        [28]   // FV26 Chill Down Pressure
        [29]   // FV26 Chill Down Current Time
        [2]   // FV26 Level Probes
        [30]   // FV26 Time since Clean
        [32]   // FV26 CIP Selected
        [32].0   // FV26 Request Channel 1 CIP
        [32].1   // FV26 Request Channel 2 CIP
        [33]   // FV26 Rotocheck
        [33].0   // FV26 Enable Rotocheck
        [33].1   // FV26 Rotocheck Fault
        [38]   // FV26 Pressure Difference Bottom-Top (psi)
        [39]   // FV26 Pressure Difference Calibration Offset
        [3]   // FV26 Top Pressure Status
        [40]   // FV26 Cropping Status 0=Not Done 1=Running 2=Done 3=Done+48hrs
        [43]   // FV26 Hours since Yeast Cropping
        [4]   // FV26 Yeast Status
        [50]   // FV26 FiltrateReturnStatus 0=Not Done 1=Running 2=Done
        [5]   // FV26 Aging Status
        [60].3   // FV26 Top Pressure Chill Down
        [6]   // FV26 Valve Routes
        [6].0   // FV26 Inlet Main to Drain Open
        [6].1   // FV26 Filling Valve Not Closed
        [6].2   // FV26 Filling Inlet Open
        [6].3   // FV26 Bypass Route Open Open
        [6].4   // FV26 Green Beer Open
        [6].5   // FV26 Yeast Removal Open
        [6].6   // FV26 Filtrate Open
        [6].7   // FV26 CIP Open
        [7]   // FV26 Top Pressure Control Actual Pressure
        [7].0   // FV26 Yeast Status Filtrate Return
        [8]   // FV26 Log Message
        [9]   // FV26 Item Fault
   FR_N27 : INT[265] := ([0] := 227, [1] := 3, [3] := 2, [5] := 4, [6] := 8, [7] := 1030, [8] := 12227, [9] := -1, [10] := 2387, [11] := 9672, [12] := 1575, [13] := 2902, [14] := 603, [15] := 1292, [16] := 891, [17] := 9083, [18] := 12, [19] := 8975, [20] := 1, [21] := 4, [22] := 1000, [23] := 50, [24] := 1050, [25] := 950, [26] := 1000, [27] := 8, [30] := 2, [33] := 1, [37] := 702, [38] := 1357, [39] := 65, [52] := 1, [60] := 4, [68] := 5311, [69] := 172, [90] := 1, [91] := 251, [92] := 841, [100] := 43, [101] := 49, [102] := 55, [103] := 13, [104] := 14, [105] := 15, [106] := 16, [107] := 17, [108] := 97, [109] := -1, [110] := -1, [111] := -1, [112] := -1, [113] := -1, [114] := -1, [115] := -1, [116] := -1, [117] := -1, [118] := -1, [119] := -1, [120] := -1, [121] := -1,
        [122] := -1, [123] := -1, [124] := -1, [125] := -1, [126] := -1, [127] := -1, [128] := -1, [129] := -1, [130] := -1, [131] := -1, [132] := -1, [133] := -1, [134] := -1, [135] := -1, [136] := -1, [137] := -1, [138] := -1, [139] := -1, [140] := -1, [141] := -1, [142] := -1, [143] := -1, [144] := -1, [145] := -1, [146] := -1, [147] := -1, [148] := -1, [149] := -1);   // FV27
        [0]   // FV27
        [100]   // FV27 Checklist Data
        [10]   // FV27 Bottom Pressure
        [11]   // FV27 Damped Level
        [12]   // FV27 Cone Radius
        [13]   // FV27 Cone Height
        [14]   // FV27 Volume (HL)
        [19]   // FV27 Height above LTX
        [1]   // FV27 Status 0=Clean,1=Fill,2=Par t,3=Ferment,4=?,5=?, 6=?,7=?,8=Emptying,9 =Dirty,10-13=CIP
        [20]   // FV27 Top Pressure Bits
        [20].2   // FV27 Top Pressure Chill Down
        [20].5   // FV27 Top Pressure Step Channel 1 CIP
        [20].6   // FV27 Top Pressure Bits Ch1 CIP Complete
        [20].7   // FV27 Top Pressure Step Channel 2 CIP
        [20].8   // FV27 Top Pressure Bits Ch2 CIP Complete
        [21]   // FV27 Top Pressure Step Flags
        [21].0   // FV27 Top Pressure Control Over Pressure
        [21].4   // FV27 Top Pressure Open Vent
        [21].5   // FV27 Top Pressure Control Open Vent Actuator
        [21].6   // FV27 Over Top Pressure Limit
        [21].8   // FV27 Top Pressure Control Over Pressure Alarm
        [22]   // FV27 Top Pressure Setpoint
        [23]   // FV27 Top Pressure Deadband
        [24]   // FV27 Top Pressure Upper Limit
        [25]   // FV27 Top Pressure Lower Limit
        [26]   // FV27 Fermenting Pressure
        [27]   // FV27 Chill Down Time
        [28]   // FV27 Chill Down Pressure
        [29]   // FV27 Chill Down Current Time
        [2]   // FV27 Level Probes
        [30]   // FV27 Time since Clean
        [32]   // FV27 CIP Selected
        [32].0   // FV27 Request Channel 1 CIP
        [32].1   // FV27 Request Channel 2 CIP
        [33]   // FV27 Rotocheck
        [33].0   // FV27 Enable Rotocheck
        [33].1   // FV27 Rotocheck Fault
        [38]   // FV27 Pressure Difference Bottom-Top (psi)
        [39]   // FV27 Pressure Difference Calibration Offset
        [3]   // FV27 Top Pressure Status
        [40]   // FV27 Cropping Status 0=Not Done 1=Running 2=Done 3=Done+48hrs
        [43]   // FV27 Hours since Yeast Cropping
        [4]   // FV27 Yeast Status
        [50]   // FV27 FiltrateReturnStatus 0=Not Done 1=Running 2=Done
        [5]   // FV27 Aging Status
        [60].3   // FV27 Top Pressure Chill Down
        [6]   // FV27 Valve Routes
        [6].0   // FV27 Inlet Main to Drain Open
        [6].1   // FV27 Filling Valve Not Closed
        [6].2   // FV27 Filling Inlet Open
        [6].3   // FV27 Bypass Route Open Open
        [6].4   // FV27 Green Beer Open
        [6].5   // FV27 Yeast Removal Open
        [6].6   // FV27 Filtrate Open
        [6].7   // FV27 CIP Open
        [7]   // FV27 Top Pressure Control Actual Pressure
        [7].0   // FV27 Yeast Status Filtrate Return
        [8]   // FV27 Log Message
        [90]   // Vent Actuations Counter
        [91]   // FV27/PTX01 FV27 top pressure minimum
        [92]   // FV27/PTX01 FV27 top pressure maximum
        [9]   // FV27 Item Fault
   FR_N28 : INT[265] := ([0] := 228, [1] := 3, [2] := 1, [3] := 4, [4] := 30, [5] := 6, [6] := 8, [7] := 1, [8] := 12228, [9] := -1, [10] := 1150, [11] := 8680, [12] := 1575, [13] := 2902, [14] := 526, [15] := 1149, [16] := 792, [17] := 8073, [18] := 12, [19] := 7977, [20] := 1, [21] := 18, [22] := 167, [24] := 167, [25] := 167, [26] := 1000, [27] := 12, [29] := 10, [30] := 23, [33] := 1, [37] := 702, [38] := 1149, [52] := 1, [60] := 16, [68] := 5228, [69] := 5228, [100] := 47, [101] := 53, [102] := 59, [103] := 27, [104] := 28, [105] := 29, [106] := 30, [107] := 31, [108] := 98, [109] := -1, [110] := -1, [111] := -1, [112] := -1, [113] := -1, [114] := -1, [115] := -1, [116] := -1, [117] := -1, [118] := -1, [119] := -1, [120] := -1, [121] := -1, [122] := -1, [123] := -1,
        [124] := -1, [125] := -1, [126] := -1, [127] := -1, [128] := -1, [129] := -1, [130] := -1, [131] := -1, [132] := -1, [133] := -1, [134] := -1, [135] := -1, [136] := -1, [137] := -1, [138] := -1, [139] := -1, [140] := -1, [141] := -1, [142] := -1, [143] := -1, [144] := -1, [145] := -1, [146] := -1, [147] := -1, [148] := -1, [149] := -1);   // FV28
        [0]   // FV28
        [100]   // FV28 Checklist Data
        [10]   // FV28 Bottom Pressure
        [11]   // FV28 Damped Level
        [12]   // FV28 Cone Radius
        [13]   // FV28 Cone Height
        [14]   // FV28 Volume (HL)
        [19]   // FV28 Height above LTX
        [1]   // FV28 Status 0=Clean,1=Fill,2=Par t,3=Ferment,4=?,5=?, 6=?,7=?,8=Emptying,9 =Dirty,10-13=CIP
        [20]   // FV28 Top Pressure Bits
        [20].2   // FV28 Top Pressure Chill Down
        [20].5   // FV28 Top Pressure Step Channel 1 CIP
        [20].6   // FV28 Top Pressure Bits Ch1 CIP Complete
        [20].7   // FV28 Top Pressure Step Channel 2 CIP
        [20].8   // FV28 Top Pressure Bits Ch2 CIP Complete
        [21]   // FV28 Top Pressure Step Flags
        [21].0   // FV28 Top Pressure Control Over Pressure
        [21].4   // FV28 Top Pressure Open Vent
        [21].5   // FV28 Top Pressure Control Open Vent Actuator
        [21].6   // FV28 Over Top Pressure Limit
        [21].8   // FV28 Top Pressure Control Over Pressure Alarm
        [22]   // FV28 Top Pressure Setpoint
        [23]   // FV28 Top Pressure Deadband
        [24]   // FV28 Top Pressure Upper Limit
        [25]   // FV28 Top Pressure Lower Limit
        [26]   // FV28 Fermenting Pressure
        [27]   // FV28 Chill Down Time
        [28]   // FV28 Chill Down Pressure
        [29]   // FV28 Chill Down Current Time
        [2]   // FV28 Level Probes
        [30]   // FV28 Time since Clean
        [32]   // FV28 CIP Selected
        [32].0   // FV28 Request Channel 1 CIP
        [32].1   // FV28 Request Channel 2 CIP
        [33]   // FV28 Rotocheck
        [33].0   // FV28 Enable Rotocheck
        [33].1   // FV28 Rotocheck Fault
        [38]   // FV28 Pressure Difference Bottom-Top (psi)
        [39]   // FV28 Pressure Difference Calibration Offset
        [3]   // FV28 Top Pressure Status
        [40]   // FV28 Cropping Status 0=Not Done 1=Running 2=Done 3=Done+48hrs
        [43]   // FV28 Hours since Yeast Cropping
        [4]   // FV28 Yeast Status
        [50]   // FV28 FiltrateReturnStatus 0=Not Done 1=Running 2=Done
        [5]   // FV28 Aging Status
        [60].3   // FV28 Top Pressure Chill Down
        [6]   // FV28 Valve Routes
        [6].0   // FV28 Inlet Main to Drain Open
        [6].1   // FV28 Filling Valve Not Closed
        [6].2   // FV28 Filling Inlet Open
        [6].3   // FV28 Bypass Route Open Open
        [6].4   // FV28 Green Beer Open
        [6].5   // FV28 Yeast Removal Open
        [6].6   // FV28 Filtrate Open
        [6].7   // FV28 CIP Open
        [7]   // FV28 Top Pressure Control Actual Pressure
        [7].0   // FV28 Yeast Status Filtrate Return
        [8]   // FV28 Log Message
        [9]   // FV28 Item Fault
   FR_N29 : INT[265] := ([0] := 229, [1] := 9, [2] := 2, [3] := 6, [4] := 2, [6] := 8, [7] := 6, [8] := 12229, [9] := -1, [10] := -1, [11] := -50, [12] := 1575, [13] := 2902, [15] := -7, [16] := -5, [17] := -51, [18] := 12, [19] := -50, [20] := 1, [21] := 33, [22] := -125, [23] := 50, [24] := -75, [25] := -175, [26] := 1000, [27] := 8, [30] := 39, [33] := 1, [37] := 702, [38] := -7, [52] := 1, [60] := 64, [69] := 5213, [100] := 46, [101] := 52, [102] := 58, [103] := 32, [104] := 33, [105] := 34, [106] := 35, [107] := 36, [108] := 99, [109] := -1, [110] := -1, [111] := -1, [112] := -1, [113] := -1, [114] := -1, [115] := -1, [116] := -1, [117] := -1, [118] := -1, [119] := -1, [120] := -1, [121] := -1, [122] := -1, [123] := -1, [124] := -1, [125] := -1, [126] := -1,
        [127] := -1, [128] := -1, [129] := -1, [130] := -1, [131] := -1, [132] := -1, [133] := -1, [134] := -1, [135] := -1, [136] := -1, [137] := -1, [138] := -1, [139] := -1, [140] := -1, [141] := -1, [142] := -1, [143] := -1, [144] := -1, [145] := -1, [146] := -1, [147] := -1, [148] := -1, [149] := -1);   // FV29
        [0]   // FV29
        [100]   // FV29 Checklist Data
        [10]   // FV29 Bottom Pressure
        [11]   // FV29 Damped Level
        [12]   // FV29 Cone Radius
        [13]   // FV29 Cone Height
        [14]   // FV29 Volume (HL)
        [19]   // FV29 Height above LTX
        [1]   // FV29 Status 0=Clean,1=Fill,2=Par t,3=Ferment,4=?,5=?, 6=?,7=?,8=Emptying,9 =Dirty,10-13=CIP
        [20]   // FV29 Top Pressure Bits
        [20].2   // FV29 Top Pressure Chill Down
        [20].5   // FV29 Top Pressure Step Channel 1 CIP
        [20].6   // FV29 Top Pressure Bits Ch1 CIP Complete
        [20].7   // FV29 Top Pressure Step Channel 2 CIP
        [20].8   // FV29 Top Pressure Bits Ch2 CIP Complete
        [21]   // FV29 Top Pressure Step Flags
        [21].0   // FV29 Top Pressure Control Over Pressure
        [21].4   // FV29 Top Pressure Open Vent
        [21].5   // FV29 Top Pressure Control Open Vent Actuator
        [21].6   // FV29 Over Top Pressure Limit
        [21].8   // FV29 Top Pressure Control Over Pressure Alarm
        [22]   // FV29 Top Pressure Setpoint
        [23]   // FV29 Top Pressure Deadband
        [24]   // FV29 Top Pressure Upper Limit
        [25]   // FV29 Top Pressure Lower Limit
        [26]   // FV29 Fermenting Pressure
        [27]   // FV29 Chill Down Time
        [28]   // FV29 Chill Down Pressure
        [29]   // FV29 Chill Down Current Time
        [2]   // FV29 Level Probes
        [30]   // FV29 Time since Clean
        [32]   // FV29 CIP Selected
        [32].0   // FV29 Request Channel 1 CIP
        [32].1   // FV29 Request Channel 2 CIP
        [33]   // FV29 Rotocheck
        [33].0   // FV29 Enable Rotocheck
        [33].1   // FV29 Rotocheck Fault
        [38]   // FV29 Pressure Difference Bottom-Top (psi)
        [39]   // FV29 Pressure Difference Calibration Offset
        [3]   // FV29 Top Pressure Status
        [40]   // FV29 Cropping Status 0=Not Done 1=Running 2=Done 3=Done+48hrs
        [43]   // FV29 Hours since Yeast Cropping
        [4]   // FV29 Yeast Status
        [50]   // FV29 FiltrateReturnStatus 0=Not Done 1=Running 2=Done
        [5]   // FV29 Aging Status
        [60].3   // FV29 Top Pressure Chill Down
        [6]   // FV29 Valve Routes
        [6].0   // FV29 Inlet Main to Drain Open
        [6].1   // FV29 Filling Valve Not Closed
        [6].2   // FV29 Filling Inlet Open
        [6].3   // FV29 Bypass Route Open Open
        [6].4   // FV29 Green Beer Open
        [6].5   // FV29 Yeast Removal Open
        [6].6   // FV29 Filtrate Open
        [6].7   // FV29 CIP Open
        [7]   // FV29 Top Pressure Control Actual Pressure
        [7].0   // FV29 Yeast Status Filtrate Return
        [8]   // FV29 Log Message
        [9]   // FV29 Item Fault
   FR_N30 : INT[265] := ([0] := 230, [1] := 9, [2] := 38, [3] := 6, [6] := 8, [7] := -5, [8] := 12230, [9] := -1, [10] := -7, [11] := 10, [12] := 1600, [13] := 2715, [15] := 1, [16] := 1, [17] := 10, [18] := 12, [19] := 10, [21] := 34, [22] := 83, [23] := 50, [24] := 133, [25] := 33, [26] := 1000, [27] := 12, [30] := 39, [33] := 1, [37] := 600, [38] := -2, [39] := -3, [52] := 1, [60] := 64, [69] := 749, [100] := 45, [101] := 51, [102] := 79, [103] := 64, [104] := 65, [105] := 66, [106] := 67, [107] := 68, [108] := 100, [109] := -1, [110] := -1, [111] := -1, [112] := -1, [113] := -1, [114] := -1, [115] := -1, [116] := -1, [117] := -1, [118] := -1, [119] := -1, [120] := -1, [121] := -1, [122] := -1, [123] := -1, [124] := -1, [125] := -1, [126] := -1, [127] := -1,
        [128] := -1, [129] := -1, [130] := -1, [131] := -1, [132] := -1, [133] := -1, [134] := -1, [135] := -1, [136] := -1, [137] := -1, [138] := -1, [139] := -1, [140] := -1, [141] := -1, [142] := -1, [143] := -1, [144] := -1, [145] := -1, [146] := -1, [147] := -1, [148] := -1, [149] := -1);   // FV30
        [0]   // FV30
        [100]   // FV30 Checklist Data
        [10]   // FV30 Bottom Pressure
        [11]   // FV30 Damped Level
        [12]   // FV30 Cone Radius
        [13]   // FV30 Cone Height
        [14]   // FV30 Volume (HL)
        [19]   // FV30 Height above LTX
        [1]   // FV30 Status 0=Clean,1=Fill,2=Par t,3=Ferment,4=?,5=?, 6=?,7=?,8=Emptying,9 =Dirty,10-13=CIP
        [20]   // FV30 Top Pressure Bits
        [20].2   // FV30 Top Pressure Chill Down
        [20].5   // FV30 Top Pressure Step Channel 1 CIP
        [20].6   // FV30 Top Pressure Bits Ch1 CIP Complete
        [20].7   // FV30 Top Pressure Step Channel 2 CIP
        [20].8   // FV30 Top Pressure Bits Ch2 CIP Complete
        [21]   // FV30 Top Pressure Step Flags
        [21].0   // FV30 Top Pressure Control Over Pressure
        [21].4   // FV30 Top Pressure Open Vent
        [21].5   // FV30 Top Pressure Control Open Vent Actuator
        [21].6   // FV30 Over Top Pressure Limit
        [21].8   // FV30 Top Pressure Control Over Pressure Alarm
        [22]   // FV30 Top Pressure Setpoint
        [23]   // FV30 Top Pressure Deadband
        [24]   // FV30 Top Pressure Upper Limit
        [25]   // FV30 Top Pressure Lower Limit
        [26]   // FV30 Fermenting Pressure
        [27]   // FV30 Chill Down Time
        [28]   // FV30 Chill Down Pressure
        [29]   // FV30 Chill Down Current Time
        [2]   // FV30 Level Probes
        [30]   // FV30 Time since Clean
        [32]   // FV30 CIP Selected
        [32].0   // FV30 Request Channel 1 CIP
        [32].1   // FV30 Request Channel 2 CIP
        [33]   // FV30 Rotocheck
        [33].0   // FV30 Enable Rotocheck
        [33].1   // FV30 Rotocheck Fault
        [38]   // FV30 Pressure Difference Bottom-Top (psi)
        [39]   // FV30 Pressure Difference Calibration Offset
        [3]   // FV30 Top Pressure Status
        [40]   // FV30 Cropping Status 0=Not Done 1=Running 2=Done 3=Done+48hrs
        [43]   // FV30 Hours since Yeast Cropping
        [4]   // FV30 Yeast Status
        [50]   // FV30 FiltrateReturnStatus 0=Not Done 1=Running 2=Done
        [5]   // FV30 Aging Status
        [60].3   // FV30 Top Pressure Chill Down
        [6]   // FV30 Valve Routes
        [6].0   // FV30 Inlet Main to Drain Open
        [6].1   // FV30 Filling Valve Not Closed
        [6].2   // FV30 Filling Inlet Open
        [6].3   // FV30 Bypass Route Open Open
        [6].4   // FV30 Green Beer Open
        [6].5   // FV30 Yeast Removal Open
        [6].6   // FV30 Filtrate Open
        [6].7   // FV30 CIP Open
        [7]   // FV30 Top Pressure Control Actual Pressure
        [7].0   // FV30 Yeast Status Filtrate Return
        [8]   // FV30 Log Message
        [9]   // FV30 Item Fault
   FR_N31 : INT[265] := ([0] := 231, [1] := 3, [3] := 4, [5] := 6, [6] := 8, [7] := -1, [8] := 13231, [9] := -1, [10] := 1143, [11] := 8392, [12] := 1600, [13] := 2715, [14] := 529, [15] := 1144, [16] := 789, [17] := 8043, [18] := 32, [19] := 7794, [21] := 17, [22] := -125, [23] := 50, [24] := -75, [25] := -175, [26] := 1000, [27] := 8, [29] := 10, [30] := 21, [33] := 1, [37] := 600, [38] := 1144, [52] := 1, [60] := 16, [68] := 5323, [69] := 172, [100] := 44, [101] := 50, [102] := 56, [103] := 69, [104] := 70, [105] := 71, [106] := 72, [107] := 73, [108] := 101, [109] := -1, [110] := -1, [111] := -1, [112] := -1, [113] := -1, [114] := -1, [115] := -1, [116] := -1, [117] := -1, [118] := -1, [119] := -1, [120] := -1, [121] := -1, [122] := -1, [123] := -1, [124] := -1, [125] := -1,
        [126] := -1, [127] := -1, [128] := -1, [129] := -1, [130] := -1, [131] := -1, [132] := -1, [133] := -1, [134] := -1, [135] := -1, [136] := -1, [137] := -1, [138] := -1, [139] := -1, [140] := -1, [141] := -1, [142] := -1, [143] := -1, [144] := -1, [145] := -1, [146] := -1, [147] := -1, [148] := -1, [149] := -1);   // FV31
        [0]   // FV31
        [100]   // FV31 Checklist Data
        [10]   // FV31 Bottom Pressure
        [11]   // FV31 Damped Level
        [12]   // FV31 Cone Radius
        [13]   // FV31 Cone Height
        [14]   // FV31 Volume (HL)
        [19]   // FV31 Height above LTX
        [1]   // FV31 Status 0=Clean,1=Fill,2=Par t,3=Ferment,4=?,5=?, 6=?,7=?,8=Emptying,9 =Dirty,10-13=CIP
        [20]   // FV31 Top Pressure Bits
        [20].2   // FV31 Top Pressure Chill Down
        [20].5   // FV31 Top Pressure Step Channel 1 CIP
        [20].6   // FV31 Top Pressure Bits Ch1 CIP Complete
        [20].7   // FV31 Top Pressure Step Channel 2 CIP
        [20].8   // FV31 Top Pressure Bits Ch2 CIP Complete
        [21]   // FV31 Top Pressure Step Flags
        [21].0   // FV31 Top Pressure Control Over Pressure
        [21].4   // FV31 Top Pressure Open Vent
        [21].5   // FV31 Top Pressure Control Open Vent Actuator
        [21].6   // FV31 Over Top Pressure Limit
        [21].8   // FV31 Top Pressure Control Over Pressure Alarm
        [22]   // FV31 Top Pressure Setpoint
        [23]   // FV31 Top Pressure Deadband
        [24]   // FV31 Top Pressure Upper Limit
        [25]   // FV31 Top Pressure Lower Limit
        [26]   // FV31 Fermenting Pressure
        [27]   // FV31 Chill Down Time
        [28]   // FV31 Chill Down Pressure
        [29]   // FV31 Chill Down Current Time
        [2]   // FV31 Level Probes
        [30]   // FV31 Time since Clean
        [32]   // FV31 CIP Selected
        [32].0   // FV31 Request Channel 1 CIP
        [32].1   // FV31 Request Channel 2 CIP
        [33]   // FV31 Rotocheck
        [33].0   // FV31 Enable Rotocheck
        [33].1   // FV31 Rotocheck Fault
        [38]   // FV31 Pressure Difference Bottom-Top (psi)
        [39]   // FV31 Pressure Difference Calibration Offset
        [3]   // FV31 Top Pressure Status
        [40]   // FV31 Cropping Status 0=Not Done 1=Running 2=Done 3=Done+48hrs
        [43]   // FV31 Hours since Yeast Cropping
        [4]   // FV31 Yeast Status
        [50]   // FV31 FiltrateReturnStatus 0=Not Done 1=Running 2=Done
        [5]   // FV31 Aging Status
        [60].3   // FV31 Top Pressure Chill Down
        [6]   // FV31 Valve Routes
        [6].0   // FV31 Inlet Main to Drain Open
        [6].1   // FV31 Filling Valve Not Closed
        [6].2   // FV31 Filling Inlet Open
        [6].3   // FV31 Bypass Route Open Open
        [6].4   // FV31 Green Beer Open
        [6].5   // FV31 Yeast Removal Open
        [6].6   // FV31 Filtrate Open
        [6].7   // FV31 CIP Open
        [7]   // FV31 Top Pressure Control Actual Pressure
        [7].0   // FV31 Yeast Status Filtrate Return
        [8]   // FV31 Log Message
        [9]   // FV31 Item Fault
   FR_N36 : INT[265];   // Original N File From SLC, No Description Available
        [1]   // Vessel Status 0=Clean,1=Filling,2= Beer,3=Packng1,4=Pac kng2,5=Packng3,6=Ven ting,7=Dirty,8=CIP
        [20].7   // Vessel Top Pressure Channel 2 CIP
        [21].4   // Vessel Top Pressure Open Vent
        [21].5   // Vessel Top Pressure Open CO2
        [2].1   // MV36/LLP01 MV36 Low level Debounced
        [32].0   // MV36 Channel 1 CIP Request
        [32].1   // MV36 Channel 2 CIP Request
        [6].0   // MV36 Inlet Main to Drain Open
        [6].1   // MV36 Inlet Main to Vessel Open
        [6].2   // MV36 Route Closed
   FR_N37 : INT[265];   // Original N File From SLC, No Description Available
        [20].5   // Vessel Top Pressure CIP
        [2].1   // MV37/LLP01 MV37 Low level Debounced
        [32].0   // MV37 Channel 1 CIP Request
        [32].1   // MV37 Channel 2 CIP Request
   FR_N46 : INT[265];   // Original N File From SLC, No Description Available
        [20].5   // Vessel Top Pressure CIP
        [2].1   // MV46/LLP01 MV46 Low level Debounced
        [32].0   // MV46 Channel 1 CIP Request
        [32].1   // MV46 Channel 2 CIP Request
   FR_N47 : INT[265];   // Original N File From SLC, No Description Available
        [20].5   // Vessel Top Pressure CIP
        [2].1   // MV47/LLP01 MV47 Low level Debounced
        [32].0   // MV47 Channel 1 CIP Request
        [32].1   // MV47 Channel 2 CIP Request
   FR_N7 : INT[265] := ([0] := 120, [10] := 31, [11] := 31, [13] := 1100, [16] := 2000);   // INTEGER
        [0]   // Register to trap a the source of an overflow error
        [10]   // Rotate Selected Vessel for Top Pressure
        [11]   // Selected Vessel for Top Pressure
        [13]   // FV26-29 Max Pressure
        [14]   // Any Vessel Over Top Pressure Limit
        [14].0   // Any Vessel Over Top Pressure Limit
        [15]   // Vent pipework mods complete
        [15].0   // Vent pipework mods complete
        [16]   // FV30-31 Max Pressure
   FR_N99 : INT[265] := ([2] := 3, [5] := 1, [7] := 1, [10] := 1, [26] := 15, [27] := 15, [28] := 15, [29] := 15, [30] := 15, [31] := 15, [100] := 1, [101] := 15, [102] := 1, [110] := 1, [111] := 15, [112] := 1, [120] := 1, [121] := 15, [122] := 1, [130] := 1, [131] := 23, [132] := 1, [133] := 1, [140] := 15, [141] := 1, [160] := 63, [170] := 1, [171] := 11, [172] := 1, [200] := 1, [202] := 1, [210] := 1, [220] := 3, [221] := 1, [240] := 1, [255] := 7);   // COMMENT Comment Lines
        [100].0   // FV Fill Status and Commands
        [101].0   // FV Fill Step Sequence Startup
        [101].1   // FV Fill Step Sequence Process
        [101].2   // FV Fill Step Sequence CIP
        [102].0   // FV Fill Outputs
        [10].0   // Communications to other PLCs
        [110].0   // Green Beer to Centrifuge Status and Commands
        [111].0   // Green Beer Step Sequence
        [111].1   // Green Beer Step Sequence Process
        [111].2   // Green Beer Step Sequence CIP
        [111].3   // Green Beer Step Sequence Held
        [111].4   // FV>MV Step Sequence Copy Data to MV Routing PLC
        [112].0   // Green Beer Outputs
        [120].0   // Yeast Cropping Status and Commands
        [121].0   // Yeast Cropping Step Sequence Startup
        [121].1   // Yeast Cropping Step Sequence Process
        [121].2   // Yeast Cropping Step Sequence CIP
        [121].3   // Yeast Cropping Step Sequence Held
        [122].0   // Yeast Cropping Outputs
        [130].0   // Filtrate Return Status and Commands
        [131].0   // Filtrate Return Step Sequence Startup
        [131].1   // Filtrate Return Step Sequence Process
        [131].2   // Filtrate Return Step Sequence CIP
        [131].4   // Filtrate Return Step Sequence Held
        [132].0   // Filtrate Return Outputs
        [133].0   // Filtrate Return Vessel Switch Box, Valve and Pump Control
        [140].0   // CIP Available Flags
        [140].1   // CIP Open Route/Complete Flags
        [140].2   // CIP Request Flags
        [140].3   // CIP Pulse Timers
        [141].0   // CIP Outputs
        [160].0   // Vessel Subroutine CIP Steps
        [160].1   // Vessel Subroutine Top Pressure Steps
        [160].2   // Vessel Top Pressure Step Sequence
        [160].3   // Vessel Subroutine Top Pressure Control
        [160].4   // Vessel Subroutine Alarms
        [160].5   // Vessel Subroutine Volume Calculation
        [170].0   // FV1-17 Yeast Cropping Status and Commands
        [171].0   // FV1-17 Yeast Cropping Step Sequence Startup
        [171].1   // FV1-17 Yeast Cropping Step Sequence Process
        [171].3   // FV1-17 Yeast Cropping Step Sequence Held
        [172].0   // FV1-17 Yeast Cropping Output
        [180].0   // FV18-25 Yeast Cropping Status and Commands
        [181].0   // FV18-25 Yeast Cropping Step Sequence Startup
        [181].1   // FV18-25 Yeast Cropping Step Sequence Process
        [181].3   // FV18-25 Yeast Cropping Step Sequence Held
        [182].0   // FV18-25 Yeast Cropping Output
        [200].0   // Analog Inputs
        [210].0   // Scale the Analog Outputs
        [221].0   // Scan a list of checkwords (File N[N160:200]:100) and enable checking and set to automatic
        [240].0   // Debounce the digital inputs
        [255].0   // Continuous Checking
        [26].0   // FV26 Inputs
        [26].1   // FV26 call vessel and plant item checklist subroutines
        [26].2   // FV26 drive outputs.
        [26].3   // FV26 Timers
        [27].0   // FV27 Inputs
        [27].1   // FV27 call vessel and plant item checklist subroutines
        [27].2   // FV27 drive outputs.
        [27].3   // FV27 Timers
        [28].0   // FV28 Inputs
        [28].1   // FV28 call vessel and plant item checklist subroutines
        [28].2   // FV28 drive outputs.
        [28].3   // FV28 Timers
        [29].0   // FV29 Inputs
        [29].1   // FV29 call vessel and plant item checklist subroutines
        [29].2   // FV29 drive outputs.
        [29].3   // FV29 Timers
        [3].0   // Simulation Code to be run in office only
        [4].0   // Simulation Code to be run in office only
        [5].0   // Initialisation Code
        [7].0   // General Code Siren, Beacon, General purpose timers
   FR_OXY_SW1 : PlantItem;   // OXY_SW1
   FR_OXY_SW1_RawInput : ALIAS FOR RIO_Rack_2:3:I.Data.28;   // FR_OXY_SW1
   FR_OXY_SW2 : PlantItem;   // OXY_SW2
   FR_OXY_SW2_RawInput : ALIAS FOR RIO_Rack_2:3:I.Data.29;   // FR_OXY_SW2
   FR_PANELESTOP : PlantItem := (CW := 2#0000_0000_0000_0100_0000_0000_0010_0001);   // PANELESTOP
   FR_PANELESTOP_RawInput : ALIAS FOR RIO_Rack_2:3:I.Data.30;   // FR_PANELESTOP
   FR_PANELESTOPDB : ALIAS FOR FR_B240[1].14;   // PanelEstop Panel emergency stop Debounced
   FR_PARAF : PlantItem := (CW := 2#0000_0000_0000_0100_0000_0000_0000_0001);   // PARAF
   FR_PARAF_RawInput : ALIAS FOR RIO_Rack_2:4:I.Data.4;   // FR_PARAF
   FR_PILZ : PlantItem := (CW := 2#0000_0000_0000_0100_0000_0000_0010_0001);   // PILZ
   FR_PILZ_RawInput : ALIAS FOR RIO_Rack_2:3:I.Data.31;   // FR_PILZ
   FR_PILZDB : ALIAS FOR FR_B240[1].15;   // Pilz Pilz healthy input Debounced
   FR_R3_SW3_1 : PlantItem;   // R3_SW3_1
   FR_R3_SW3_1_RawInput : ALIAS FOR RIO_Rack_2:4:I.Data.14;   // FR_R3_SW3_1 FR_N14[109].1
   FR_R3_SW3_2 : PlantItem := (CW := 2#0000_0000_0000_0100_0000_0000_0000_0001);   // R3_SW3_2
   FR_R3_SW3_2_RawInput : ALIAS FOR RIO_Rack_2:4:I.Data.10;   // FR_R3_SW3_2 FR_N14[109].0
   FR_R3_SW3_3 : PlantItem := (CW := 2#0000_0000_0000_0100_0000_0000_0000_0001);   // R3_SW3_3
   FR_R3_SW3_3_RawInput : ALIAS FOR RIO_Rack_2:3:I.Data.14;   // FR_R3_SW3_3 FR_N14[109].2
   FR_SFile : INT[255] := ([4] := -4134, [37] := 2020, [38] := 6, [39] := 22, [40] := 13, [41] := 9, [42] := 51, [53] := 3);   // SLC Equivalent System File, So Original Code Can Remain
        [1].15   // First Scan Flag
        [37]   // Clock Calendar Year
        [40]   // Clock Calendar Hours
        [41]   // Clock Calendar Minutes
        [42]   // Clock Calendar Minute
        [53]   // Calendar Day 1 = Monday
   FR_T101 : TIMER[255] := ([0].PRE := 15000, [1].PRE := 10000, [2].PRE := 3000, [10].PRE := 3000, [11].PRE := 3000, [12].PRE := 3000, [13].PRE := 3000, [14].PRE := 3000, [15].PRE := 3000, [16].PRE := 3000);   // FV FILLING
        [0]   // FV_Fill STEP Command Data Check
        [10]   // FV_Fill Cancel Prompt
        [11]   // FV_Fill STEP SCADA Prompts Beer Transfer Complete
        [1]   // Delay before O2 Valve Alarm
        [2]   // FV_Fill SCADA Prompts Abort Delay
   FR_T111 : TIMER[255] := ([0].PRE := 30000, [1].PRE := 60000, [2].PRE := 3000, [5].PRE := 3000, [6].PRE := 3000, [7].PRE := 3000, [8].PRE := 3000, [10].PRE := 3000, [11].PRE := 3000);   // GREEN BEER
        [0]   // Green Beer Wait for SCADA Data
        [10]   // Green Beer PROMPTS Cancel
        [11]   // Green Beer STEP SCADA Prompts Beer Transfer Complete
        [1]   // Green Beer STEP Water Chase
        [2]   // Green Beer SCADA Prompt Abort
        [5]   // Green Beer STEP SCADA Prompts Extend Transfer
        [6]   // Green Beer STEP SCADA Prompts Flush Main
        [7]   // Green Beer STEP SCADA Prompts End Transfer
        [8]   // Green Beer STEP SCADA Prompts End Flush
   FR_T121 : TIMER[255] := ([0].PRE := 30000, [2].PRE := 3000, [4].PRE := 60000, [5].PRE := 120000, [6].PRE := 1200000, [7].PRE := 35000, [9].PRE := 3000, [10].PRE := 3000, [11].PRE := 3000, [12].PRE := 3000, [12].ACC := 3000, [12].EN := 1, [12].DN := 1, [13].PRE := 3000, [13].ACC := 3000, [13].EN := 1, [13].DN := 1, [14].PRE := 3000, [14].ACC := 3000, [14].EN := 1, [14].DN := 1, [15].PRE := 3000, [15].ACC := 3001, [15].EN := 1, [15].DN := 1, [16].PRE := 3000, [16].ACC := 3000, [16].EN := 1, [16].DN := 1, [17].PRE := 3000, [17].ACC := 3001, [17].EN := 1, [17].DN := 1);   // YEAST CROP
        [0]   // Yeast Cropping FV26-31 Command Data Check
        [10]   // Yeast Cropping FV26-31 SCADA Prompts Cancel Delay
        [12]   // FV26-31 Channel 1 CIP Delay after Clean to check if Complete
        [13]   // FV1-17 Channel 1 CIP Delay after Clean to check if Complete
        [14]   // FV18-25 Channel 1 CIP Delay after Clean to check if Complete
        [15]   // FV26-31 Channel 2 CIP Delay after Clean to check if Complete
        [16]   // FV1-17 Channel 2 CIP Delay after Clean to check if Complete
        [17]   // FV18-25 Channel 2 CIP Delay after Clean to check if Complete
        [2]   // Yeast Cropping FV26-31 SCADA Prompts Abort Delay
        [4]   // Yeast Cropping FV26-31 Minimum Speed Duration
        [5]   // Yeast Cropping FV26-31 Ramp Up Duration
        [6]   // Yeast Cropping FV26-31 Maximum Speed Duration
        [7]   // Yeast Cropping FV26-31 Flush
   FR_T131 : TIMER[255] := ([0].PRE := 30000, [1].PRE := 30000, [2].PRE := 3000, [3].PRE := 10000, [3].ACC := 10000, [3].DN := 1, [10].PRE := 3000, [11].PRE := 3000);   // FILTRATE
        [0]   // Filtrate Return STEP Command Data Check
   FR_T141 : TIMER[255];   // CIP
   FR_T144 : TIMER[255] := ([0].PRE := 300000, [0].ACC := 24450, [0].EN := 1, [0].TT := 1, [1].PRE := 5000, [1].ACC := 5000, [1].EN := 1, [1].DN := 1, [2].PRE := 5000, [2].ACC := 5001, [2].EN := 1, [2].DN := 1, [3].PRE := 5000, [3].ACC := 5001, [3].EN := 1, [3].DN := 1, [4].PRE := 5000, [4].ACC := 5001, [4].EN := 1, [4].DN := 1, [5].PRE := 5000, [5].ACC := 4448, [5].EN := 1, [5].TT := 1, [6].PRE := 2000, [7].PRE := 5000, [8].PRE := 5000, [9].PRE := 5000, [10].PRE := 2000, [11].PRE := 2000, [12].PRE := 2000, [13].PRE := 2000, [14].PRE := 2000, [15].PRE := 2000);   // CIP
        [0]   // CIP Pulse Retrigger
        [10]   // FV26 CIP Burst Starting
        [11]   // FV27 CIP Burst Starting
        [12]   // FV28 CIP Burst Starting
        [13]   // FV29 CIP Burst Starting
        [14]   // FV30 CIP Burst Starting
        [15]   // FV31 CIP Burst Starting
        [1]   // CIP Pulse 1
        [2]   // CIP Pulse 2
        [3]   // CIP Pulse 3
        [4]   // CIP Pulse 4
        [5]   // CIP Pulse 5
        [6]   // CIP Pulse 6
        [7]   // CIP Pulse 7
        [8]   // CIP Pulse 8
        [9]   // CIP Pulse 9
   FR_T19 : TIMER[255] := ([0].PRE := 20000, [0].ACC := 417, [0].EN := 1, [0].TT := 1, [1].PRE := 20000, [2].PRE := 20000, [2].ACC := 1427, [2].EN := 1, [2].TT := 1, [3].PRE := 20000, [4].PRE := 20000, [5].PRE := 20000, [5].ACC := 417, [5].EN := 1, [5].TT := 1);   // HEARTBEAT Heartbeat Timers
        [0]   // MV_Routing_Unit Heartbeat Stuck Off
        [1]   // MV_Routing_Unit Heartbeat Stuck On
        [2]   // FV_Aging PLC Heartbeat Stuck Off
        [3]   // FV_Aging PLC Heartbeat Stuck On
        [4]   // MVFV CIP PLC Heartbeat Stuck Off
        [5]   // MVFV CIP PLC Heartbeat Stuck On
   FR_T242 : TIMER[255] := ([0].PRE := 5000, [1].PRE := 5000, [2].PRE := 5000, [3].PRE := 5000, [4].PRE := 5000, [4].ACC := 5000, [4].EN := 1, [4].DN := 1, [5].PRE := 5000, [6].PRE := 5000, [7].PRE := 5000, [7].ACC := 5000, [7].EN := 1, [7].DN := 1, [8].PRE := 5000, [9].PRE := 5000, [9].ACC := 5001, [9].EN := 1, [9].DN := 1, [10].PRE := 5000, [11].PRE := 5000, [12].PRE := 5000, [12].ACC := 5000, [12].EN := 1, [12].DN := 1, [13].PRE := 5000, [13].ACC := 5000, [13].EN := 1, [13].DN := 1, [20].PRE := 5000, [21].PRE := 5000, [22].PRE := 5000, [23].PRE := 5000, [24].PRE := 5000);   // DEBOUNCE
        [0]   // FV26/HLP01 FV26 High Level Timer
        [10]   // FV31/LLP01 FV31 High Level Timer
        [11]   // FV31/HLP01 FV31 Low Level Timer
        [12]   // VB4/LP01 VB4 Vent level Timer
        [13]   // FRV1/LP01 Filtrate Return Vess Level Probe Timer
        [14]   // 0 0 Timer
        [15]   // 0 0 Timer
        [16]   // 0 0 Timer
        [17]   // 0 0 Timer
        [18]   // 0 0 Timer
        [19]   // 0 0 Timer
        [1]   // FV26/LLP01 FV26 Low Level Timer
        [20]   // 0 0 Timer
        [21]   // 0 0 Timer
        [22]   // 0 0 Timer
        [23]   // 0 0 Timer
        [24]   // 0 0 Timer
        [25]   // 0 0 Timer
        [26]   // 0 0 Timer
        [27]   // 0 0 Timer
        [28]   // 0 0 Timer
        [29]   // 0 0 Timer
        [2]   // FV27/HLP01 FV27 High Level Timer
        [30]   // PanelEstop Panel emergency stop Timer
        [31]   // Pilz Pilz healthy input Timer
        [3]   // FV27/LLP01 FV27 Low Level Timer
        [4]   // FV28/HLP01 FV28 High Level Timer
        [5]   // FV28/LLP01 FV28 Low Level Timer
        [6]   // FV29/HLP01 FV29 High Level Timer
        [7]   // FV29/LLP01 FV29 Low Level Timer
        [8]   // FV30/LLP01 FV30 High Level Timer
        [9]   // FV30/HLP01 FV30 Low Level Timer
   FR_T243 : TIMER[255] := ([0].PRE := 5000, [0].ACC := 5001, [0].EN := 1, [0].DN := 1, [1].PRE := 5000, [1].ACC := 5000, [1].EN := 1, [1].DN := 1, [2].PRE := 5000, [2].ACC := 5001, [2].EN := 1, [2].DN := 1, [3].PRE := 5000, [3].ACC := 5001, [3].EN := 1, [3].DN := 1, [4].PRE := 5000, [5].PRE := 5000, [5].ACC := 5000, [5].EN := 1, [5].DN := 1, [6].PRE := 5000, [6].ACC := 5001, [6].EN := 1, [6].DN := 1, [7].PRE := 5000, [8].PRE := 5000, [8].ACC := 5000, [8].EN := 1, [8].DN := 1, [9].PRE := 5000, [10].PRE := 5000, [10].ACC := 5000, [10].EN := 1, [10].DN := 1, [11].PRE := 5000, [11].ACC := 5000, [11].EN := 1, [11].DN := 1, [12].PRE := 1000, [13].PRE := 5000, [20].PRE := 5000, [21].PRE := 5000, [22].PRE := 5000, [23].PRE := 5000, [24].PRE := 5000);   // DEBOUNCE
        [0]   // FV26/HLP01 FV26 High Level Timer
        [10]   // FV31/LLP01 FV31 High Level Timer
        [11]   // FV31/HLP01 FV31 Low Level Timer
        [12]   // VB4/LP01 VB4 Vent level Timer
        [13]   // FRV1/LP01 Filtrate Return Vess Level Probe Timer
        [14]   // 0 0 Timer
        [15]   // 0 0 Timer
        [16]   // 0 0 Timer
        [17]   // 0 0 Timer
        [18]   // 0 0 Timer
        [19]   // 0 0 Timer
        [1]   // FV26/LLP01 FV26 Low Level Timer
        [20]   // 0 0 Timer
        [21]   // 0 0 Timer
        [22]   // 0 0 Timer
        [23]   // 0 0 Timer
        [24]   // 0 0 Timer
        [25]   // 0 0 Timer
        [26]   // 0 0 Timer
        [27]   // 0 0 Timer
        [28]   // 0 0 Timer
        [29]   // 0 0 Timer
        [2]   // FV27/HLP01 FV27 High Level Timer
        [30]   // PanelEstop Panel emergency stop Timer
        [31]   // Pilz Pilz healthy input Timer
        [3]   // FV27/LLP01 FV27 Low Level Timer
        [4]   // FV28/HLP01 FV28 High Level Timer
        [5]   // FV28/LLP01 FV28 Low Level Timer
        [6]   // FV29/HLP01 FV29 High Level Timer
        [7]   // FV29/LLP01 FV29 Low Level Timer
        [8]   // FV30/LLP01 FV30 High Level Timer
        [9]   // FV30/HLP01 FV30 Low Level Timer
   FR_T244 : TIMER[255] := ([0].PRE := 10000, [1].PRE := 10000, [2].PRE := 2000);   // CHECKWORD Checkword Timers
        [0]   // Valve Cycling Timer A
        [1]   // Valve Cycling Timer B
        [2]   // Checking Timebase
   FR_T4 : TIMER[255] := ([0].PRE := 1000, [0].ACC := 39, [0].EN := 1, [0].TT := 1, [1].PRE := 6000, [1].ACC := 2515, [1].EN := 1, [1].TT := 1, [2].PRE := 60000, [2].ACC := 53139, [2].EN := 1, [2].TT := 1, [3].PRE := 1000, [3].ACC := 348, [3].EN := 1, [3].TT := 1, [4].PRE := 1000, [5].PRE := 6000, [5].ACC := 3113, [5].EN := 1, [5].TT := 1, [6].PRE := 6000, [7].PRE := 60000, [7].ACC := 23312, [7].EN := 1, [7].TT := 1, [8].PRE := 60000, [10].PRE := 327670, [11].PRE := 20000, [11].ACC := 4824, [11].EN := 1, [11].TT := 1, [12].PRE := 2000, [12].ACC := 2000, [12].EN := 1, [12].DN := 1, [13].PRE := 1000, [14].PRE := 1000, [15].PRE := 1000, [16].PRE := 1000, [20].PRE := 30000, [21].PRE := 30000, [22].PRE := 30000, [23].PRE := 30000, [30].PRE := 10000, [31].PRE := 10000, [35].PRE := 35000, [36].PRE := 20000, [37].PRE := 5000, [38].PRE := 15000, [38].ACC := 15000, [38].EN := 1, [38].DN := 1, [39].PRE := 5000, [40].PRE := 15000, [41].PRE := 25000);   // TIMER
        [0]   // 1s Pulse
        [0].DN   // 1s pulse
        [10]   // Vent Actuations Timer
        [11]   // Rotate Selected Vessel for Top Pressure
        [12]   // Selected Vessel for Top Pressure
        [13]   // FV26 CIP Vent Pulse
        [14]   // FV27 CIP Vent Pulse
        [15]   // FV28 CIP Vent Pulse
        [16]   // FV29 CIP Vent Pulse
        [17]   // FV30 CIP Vent Pulse
        [18]   // FV31 CIP Vent Pulse
        [1]   // 6s Pulse
        [20]   // FV26 Filtrate Return Drain Gas Main
        [21]   // FV27 Filtrate Return Drain Gas Main
        [22]   // FV28 Filtrate Return Drain Gas Main
        [23]   // FV29 Filtrate Return Drain Gas Main
        [24]   // FV30 Filtrate Return Drain Gas Main
        [25]   // FV31 Filtrate Return Drain Gas Main
        [2]   // 60s Pulse
        [30]   // GEA watchdog On
        [31]   // GEA watchdog Off
        [35]   // YEAST COLLECTION H/L TIMER
        [36]   // YEAST COLLECTION RINSE START DELAY
        [37]   // YEAST COLLECTION L/L OFF
        [37].DN   // YEAST COLLECTION L/L OFF
        [38]   // YEAST COLLECTION LL START TIMER
        [38].DN   // YEAST COLLECTION LL START TIMER
        [39]   // DE-FOAMER RINSE OUT RUN TIMER
        [39].TT   // RUNNING SIGNAL FOR DE-FOAMER PUMP
        [39].DN   // DE-FOAMER TIMER DONE
        [3]   // 1s Square
        [40]   // RINSE SOL OFF DELAY
        [4]   // 1s Inverted Square
        [5]   // 6s Square
        [6]   // 6s Inverted Square
        [7]   // 60s Square
        [8]   // 60s Inverted Square
   FR_T50 : TIMER[52] := ([0].PRE := 3600000, [1].PRE := 3600000, [2].PRE := 3600000, [3].PRE := 3600000, [4].PRE := 3600000, [5].PRE := 3600000, [6].PRE := 90000, [7].PRE := 90000, [8].PRE := 90000, [9].PRE := 90000, [10].PRE := 90000, [11].PRE := 90000, [12].PRE := 5000, [13].PRE := 5000, [14].PRE := 5000, [15].PRE := 5000, [16].PRE := 5000, [17].PRE := 5000, [26].PRE := 3600000, [27].PRE := 3600000, [28].PRE := 3600000, [29].PRE := 3600000, [30].PRE := 3600000, [31].PRE := 3600000);
        [0]   // FV26 Time since Clean
        [10]   // FV30 Rotocheck Input On
        [11]   // FV31 Rotocheck Input On
        [12]   // FV26 Rotocheck Input On
        [13]   // FV27 Rotocheck Input Off
        [14]   // FV28 Rotocheck Input Off
        [15]   // FV29 Rotocheck Input Off
        [16]   // FV30 Rotocheck Input Off
        [17]   // FV31 Rotocheck Input Off
        [1]   // FV27 Time since Clean
        [26]   // FV26 Post Chill Down Timer
        [27]   // FV27 Post Chill Down Timer
        [28]   // FV28 Post Chill Down Timer
        [29]   // FV29 Post Chill Down Timer
        [2]   // FV28 Time since Clean
        [30]   // FV30 Post Chill Down Timer
        [31]   // FV31 Post Chill Down Timer
        [3]   // FV29 Time since Clean
        [4]   // FV30 Time since Clean
        [5]   // FV31 Time since Clean
        [6]   // FV26 Rotocheck Input Off
        [7]   // FV27 Rotocheck Input On
        [8]   // FV28 Rotocheck Input On
        [9]   // FV29 Rotocheck Input On
   FR_T51 : TIMER[52] := ([26].PRE := 3600000, [27].PRE := 3600000, [28].PRE := 3600000, [29].PRE := 3600000, [30].PRE := 3600000, [31].PRE := 3600000);
        [26]   // FV26 Post Yeast Cropping Timer
        [27]   // FV27 Post Yeast Cropping Timer
        [28]   // FV28 Post Yeast Cropping Timer
        [29]   // FV29 Post Yeast Cropping Timer
        [30]   // FV30 Post Yeast Cropping Timer
        [31]   // FV31 Post Yeast Cropping Timer
   FR_T52 : TIMER[52] := ([26].PRE := 180000, [26].ACC := 130290, [26].EN := 1, [26].TT := 1, [27].PRE := 180000, [28].PRE := 180000, [29].PRE := 180000, [30].PRE := 180000, [31].PRE := 180000, [31].ACC := 13218, [31].EN := 1, [31].TT := 1);
        [26]   // FV26 Top Pressure Control Over Pressure Alarm
        [27]   // FV27 Top Pressure Control Over Pressure Alarm
        [28]   // FV28 Top Pressure Control Over Pressure Alarm
        [29]   // FV29 Top Pressure Control Over Pressure Alarm
        [30]   // FV30 Top Pressure Control Over Pressure Alarm
        [31]   // FV31 Top Pressure Control Over Pressure Alarm
   FR_T53 : TIMER[52] := ([26].PRE := 30000, [27].PRE := 30000, [28].PRE := 30000, [29].PRE := 30000, [30].PRE := 30000, [31].PRE := 30000);
        [26]   // FV26 CIP Drain Down
        [27]   // FV27 CIP Drain Down
        [28]   // FV28 CIP Drain Down
        [29]   // FV29 CIP Drain Down
        [30]   // FV30 CIP Drain Down
        [31]   // FV31 CIP Drain Down
   FR_temp_real : REAL;
   fr_test_start_green_beer : BOOL;
   fr_test_start_yeast_cropping : BOOL;
   FR_to_data_file : DINT := 31;
   FR_to_data_offset : DINT := 70;
   FR_value_to_set : DINT := 160;
   FR_VB1_AV01 : PlantItem := (CW := 2#0000_0000_0000_0000_0000_0000_0011_0000, CheckTime := 10, CheckTimer := 10);   // VB1_AV01
   FR_VB1_AV01_ALARM : ALARM_DIGITAL;
   FR_VB1_AV01_C : ALIAS FOR RIO_Rack_2:6:I.Data.6;
   FR_VB1_AV01_DR : ALIAS FOR RIO_Rack_2:5:O.Data.18;
   FR_VB1_AV01_O : ALIAS FOR RIO_Rack_2:6:I.Data.2;
   FR_VB1_AV02 : PlantItem := (CW := 2#0000_0000_0000_0000_0000_0000_0001_0000, CheckTime := 10, CheckTimer := 10);   // VB1_AV02
   FR_VB1_AV02_ALARM : ALARM_DIGITAL;
   FR_VB1_AV02_C : ALIAS FOR RIO_Rack_2:6:I.Data.7;
   FR_VB1_AV02_DR : ALIAS FOR RIO_Rack_2:5:O.Data.19;
   FR_VB1_AV02_O : ALIAS FOR RIO_Rack_2:6:I.Data.3;
   FR_VB1_AV03 : PlantItem := (CW := 2#0000_0000_0000_0000_0000_0000_0001_0000, CheckTime := 10, CheckTimer := 10);   // VB1_AV03
   FR_VB1_AV03_ALARM : ALARM_DIGITAL;
   FR_VB1_AV03_C : ALIAS FOR RIO_Rack_2:6:I.Data.12;
   FR_VB1_AV03_DR : ALIAS FOR RIO_Rack_2:5:O.Data.20;
   FR_VB1_AV03_O : ALIAS FOR RIO_Rack_2:6:I.Data.8;
   FR_VB1_AV04 : PlantItem := (CW := 2#0000_0000_0000_0000_0000_0000_0001_0000, CheckTime := 10, CheckTimer := 10);   // VB1_AV04
   FR_VB1_AV04_ALARM : ALARM_DIGITAL;
   FR_VB1_AV04_C : ALIAS FOR RIO_Rack_2:6:I.Data.13;
   FR_VB1_AV04_DR : ALIAS FOR RIO_Rack_2:5:O.Data.21;
   FR_VB1_AV04_O : ALIAS FOR RIO_Rack_2:6:I.Data.9;
   FR_VB1_AV05 : PlantItem := (CW := 2#0000_0000_0000_0000_0000_0000_0001_0000, CheckTime := 10, CheckTimer := 10);   // VB1_AV05
   FR_VB1_AV05_ALARM : ALARM_DIGITAL;
   FR_VB1_AV05_C : ALIAS FOR RIO_Rack_2:6:I.Data.14;
   FR_VB1_AV05_DR : ALIAS FOR RIO_Rack_2:5:O.Data.22;
   FR_VB1_AV05_O : ALIAS FOR RIO_Rack_2:6:I.Data.10;
   FR_VB1_AV06 : PlantItem := (CW := 2#0000_0000_0000_0000_0000_0000_0001_0000, CheckTime := 10, CheckTimer := 10);   // VB1_AV06
   FR_VB1_AV06_ALARM : ALARM_DIGITAL;
   FR_VB1_AV06_C : ALIAS FOR RIO_Rack_2:6:I.Data.15;
   FR_VB1_AV06_DR : ALIAS FOR RIO_Rack_2:5:O.Data.23;
   FR_VB1_AV06_O : ALIAS FOR RIO_Rack_2:6:I.Data.11;
   FR_VB1_AV07 : PlantItem := (CW := 2#0000_0000_0000_0000_0000_0000_0001_0000, CheckTime := 10, CheckTimer := 10);   // VB1_AV07
   FR_VB1_AV07_ALARM : ALARM_DIGITAL;
   FR_VB1_AV07_C : ALIAS FOR RIO_Rack_2:6:I.Data.20;
   FR_VB1_AV07_DR : ALIAS FOR RIO_Rack_2:5:O.Data.24;
   FR_VB1_AV07_O : ALIAS FOR RIO_Rack_2:6:I.Data.16;
   FR_VB1_AV08 : PlantItem := (CW := 2#0000_0000_0000_0000_0000_0000_0000_1000, CheckTime := 10, CheckTimer := 10);   // VB1_AV08
   FR_VB1_AV08_ALARM : ALARM_DIGITAL;
   FR_VB1_AV08_C : ALIAS FOR RIO_Rack_2:6:I.Data.21;
   FR_VB1_AV08_O : ALIAS FOR RIO_Rack_2:6:I.Data.17;
   FR_VB1_AV08_RDR : ALIAS FOR RIO_Rack_2:5:O.Data.25;
   FR_VB1_AV09 : PlantItem := (CW := 2#0000_0000_0000_0000_0000_0000_0001_0000, CheckTime := 10, CheckTimer := 10);   // VB1_AV09
   FR_VB1_AV09_ALARM : ALARM_DIGITAL;
   FR_VB1_AV09_C : ALIAS FOR RIO_Rack_2:6:I.Data.22;
   FR_VB1_AV09_DR : ALIAS FOR RIO_Rack_2:5:O.Data.26;
   FR_VB1_AV09_O : ALIAS FOR RIO_Rack_2:6:I.Data.18;
   FR_VB2_AV01 : PlantItem := (CW := 2#0000_0000_0000_0000_0000_0000_0001_0000, CheckTime := 10, CheckTimer := 10);   // VB2_AV01
   FR_VB2_AV01_ALARM : ALARM_DIGITAL;
   FR_VB2_AV01_C : ALIAS FOR RIO_Rack_2:7:I.Data.13;
   FR_VB2_AV01_DR : ALIAS FOR RIO_Rack_2:8:O.Data.5;
   FR_VB2_AV01_O : ALIAS FOR RIO_Rack_2:7:I.Data.9;
   FR_VB2_AV02 : PlantItem := (CW := 2#0000_0000_0000_0000_0000_0000_0001_0000, CheckTime := 10, CheckTimer := 10);   // VB2_AV02
   FR_VB2_AV02_ALARM : ALARM_DIGITAL;
   FR_VB2_AV02_C : ALIAS FOR RIO_Rack_2:7:I.Data.14;
   FR_VB2_AV02_DR : ALIAS FOR RIO_Rack_2:8:O.Data.6;
   FR_VB2_AV02_O : ALIAS FOR RIO_Rack_2:7:I.Data.10;
   FR_VB2_AV03 : PlantItem := (CW := 2#0000_0000_0000_0000_0000_0000_0001_0000, CheckTime := 10, CheckTimer := 10);   // VB2_AV03
   FR_VB2_AV03_ALARM : ALARM_DIGITAL;
   FR_VB2_AV03_C : ALIAS FOR RIO_Rack_2:7:I.Data.15;
   FR_VB2_AV03_DR : ALIAS FOR RIO_Rack_2:8:O.Data.7;
   FR_VB2_AV03_O : ALIAS FOR RIO_Rack_2:7:I.Data.11;
   FR_VB2_AV04 : PlantItem := (CW := 2#0000_0000_0000_0000_0000_0000_0000_1000, CheckTime := 10, CheckTimer := 10);   // VB2_AV04
   FR_VB2_AV04_ALARM : ALARM_DIGITAL;
   FR_VB2_AV04_C : ALIAS FOR RIO_Rack_2:7:I.Data.20;
   FR_VB2_AV04_O : ALIAS FOR RIO_Rack_2:7:I.Data.16;
   FR_VB2_AV04_RDR : ALIAS FOR RIO_Rack_2:8:O.Data.8;
   FR_VB2_AV05 : PlantItem := (CW := 2#0000_0000_0000_0000_0000_0000_0001_0000, CheckTime := 10, CheckTimer := 10);   // VB2_AV05
   FR_VB2_AV05_ALARM : ALARM_DIGITAL;
   FR_VB2_AV05_C : ALIAS FOR RIO_Rack_2:7:I.Data.21;
   FR_VB2_AV05_DR : ALIAS FOR RIO_Rack_2:8:O.Data.9;
   FR_VB2_AV05_O : ALIAS FOR RIO_Rack_2:7:I.Data.17;
   FR_VB3_AV01 : PlantItem := (CW := 2#0000_0000_0000_0000_0000_0000_0001_0000, CheckTime := 10, CheckTimer := 10);   // VB3_AV01
   FR_VB3_AV01_ALARM : ALARM_DIGITAL;
   FR_VB3_AV01_C : ALIAS FOR RIO_Rack_2:10:I.Data.22;
   FR_VB3_AV01_DR : ALIAS FOR RIO_Rack_2:11:O.Data.10;
   FR_VB3_AV01_O : ALIAS FOR RIO_Rack_2:10:I.Data.18;
   FR_VB3_AV02 : PlantItem := (CW := 2#0000_0000_0000_0000_0000_0000_0001_0000, CheckTime := 10, CheckTimer := 10);   // VB3_AV02
   FR_VB3_AV02_ALARM : ALARM_DIGITAL;
   FR_VB3_AV02_C : ALIAS FOR RIO_Rack_2:10:I.Data.23;
   FR_VB3_AV02_DR : ALIAS FOR RIO_Rack_2:11:O.Data.11;
   FR_VB3_AV02_O : ALIAS FOR RIO_Rack_2:10:I.Data.19;
   FR_VB3_AV03 : PlantItem := (CW := 2#0000_0000_0000_0000_0000_0000_0001_0000, CheckTime := 10, CheckTimer := 10);   // VB3_AV03
   FR_VB3_AV03_ALARM : ALARM_DIGITAL;
   FR_VB3_AV03_C : ALIAS FOR RIO_Rack_2:10:I.Data.28;
   FR_VB3_AV03_DR : ALIAS FOR RIO_Rack_2:11:O.Data.12;
   FR_VB3_AV03_O : ALIAS FOR RIO_Rack_2:10:I.Data.24;
   FR_VB3_AV04 : PlantItem := (CW := 2#0000_0000_0000_0000_0000_0000_0000_1000, CheckTime := 10, CheckTimer := 10);   // VB3_AV04
   FR_VB3_AV04_ALARM : ALARM_DIGITAL;
   FR_VB3_AV04_C : ALIAS FOR RIO_Rack_2:10:I.Data.29;
   FR_VB3_AV04_O : ALIAS FOR RIO_Rack_2:10:I.Data.25;
   FR_VB3_AV04_RDR : ALIAS FOR RIO_Rack_2:11:O.Data.13;
   FR_VB3_AV05 : PlantItem := (CW := 2#0000_0000_0000_0000_0000_0000_0001_0000, CheckTime := 10, CheckTimer := 10);   // VB3_AV05
